   MCC1201_rgtDiagModule_HMI : GP_NetworkDiag_v1[50] := ([0].xFaulted := 1, [0].dEntryStatus := 16#0000_1000, [0].dFaultCode := 16#0000_0115, [0].dInstance := 16#0000_fdae, [1].xFaulted := 1, [1].dEntryStatus := 16#0000_1000, [1].dFaultCode := 16#0000_0115, [1].dInstance := 16#0000_3b39, [2].xConnected := 1, [2].dEntryStatus := 16#0000_4000, [2].dInstance := 16#0000_a3f5, [3].xConnected := 1, [3].dEntryStatus := 16#0000_7000, [3].dInstance := 16#0000_f5ac, [4].xConnected := 1, [4].dEntryStatus := 16#0000_7000, [4].dInstance := 16#0000_87af, [5].xFaulted := 1, [5].dEntryStatus := 16#0000_3000, [5].dFaultCode := 16#0000_0204, [5].dInstance := 16#0000_ac4a, [6].xFaulted := 1, [6].dEntryStatus := 16#0000_3000, [6].dFaultCode := 16#0000_0204, [6].dInstance := 16#0000_482b, [7].xFaulted := 1, [7].dEntryStatus := 16#0000_3000, [7].dFaultCode := 16#0000_0204, [7].dInstance := 16#0000_9886, [8].xFaulted := 1, [8].dEntryStatus := 16#0000_3000, [8].dFaultCode := 16#0000_0204, [8].dInstance := 16#0000_f085, [9].xFaulted := 1, [9].dEntryStatus := 16#0000_3000, [9].dFaultCode := 16#0000_0204, [9].dInstance := 16#0000_4058, [10].xFaulted := 1, [10].dEntryStatus := 16#0000_1000, [10].dFaultCode := 16#0000_0204, [10].dInstance := 16#0000_406f, [11].xFaulted := 1, [11].dEntryStatus := 16#0000_3000, [11].dFaultCode := 16#0000_0204, [11].dInstance := 16#0000_dc7a, [12].xConnected := 1, [12].dEntryStatus := 16#0000_4000, [12].dInstance := 16#0000_6808, [13].xConnected := 1, [13].dEntryStatus := 16#0000_4000, [13].dInstance := 16#0000_1271, [14].xConnected := 1, [14].dEntryStatus := 16#0000_4000, [14].dInstance := 16#0000_7aa0, [15].xConnected := 1, [15].dEntryStatus := 16#0000_4000, [15].dInstance := 16#0000_c3a3, [16].xConnected := 1, [16].dEntryStatus := 16#0000_4000, [16].dInstance := 16#0000_3650,
        [17].xConnected := 1, [17].dEntryStatus := 16#0000_4000, [17].dInstance := 16#0000_c67a, [18].xConnected := 1, [18].dEntryStatus := 16#0000_4000, [18].dInstance := 16#0000_cbaa, [19].xConnected := 1, [19].dEntryStatus := 16#0000_4000, [19].dInstance := 16#0000_7c6b, [20].xConnected := 1, [20].dEntryStatus := 16#0000_4000, [20].dInstance := 16#0000_b922, [21].xConnected := 1, [21].dEntryStatus := 16#0000_4000, [21].dInstance := 16#0000_0b41, [22].xConnected := 1, [22].dEntryStatus := 16#0000_4000, [22].dInstance := 16#0000_0a60, [23].xConnected := 1, [23].dEntryStatus := 16#0000_4000, [23].dInstance := 16#0000_ec63, [24].xConnected := 1, [24].dEntryStatus := 16#0000_4000, [24].dInstance := 16#0000_c43a, [25].xConnected := 1, [25].dEntryStatus := 16#0000_4000, [25].dInstance := 16#0000_ef15, [26].xConnected := 1, [26].dEntryStatus := 16#0000_4000, [26].dInstance := 16#0000_5364, [27].xConnected := 1, [27].dEntryStatus := 16#0000_4000, [27].dInstance := 16#0000_03d7, [28].xConnected := 1, [28].dEntryStatus := 16#0000_4000, [28].dInstance := 16#0000_365e, [29].xConnected := 1, [29].dEntryStatus := 16#0000_4000, [29].dInstance := 16#0000_bf29, [30].xConnected := 1, [30].dEntryStatus := 16#0000_4000, [30].dInstance := 16#0000_7fa8, [31].xConnected := 1, [31].dEntryStatus := 16#0000_4000, [31].dInstance := 16#0000_798b, [32].xConnected := 1, [32].dEntryStatus := 16#0000_4000, [32].dInstance := 16#0000_75c2, [33].xConnected := 1, [33].dEntryStatus := 16#0000_4000, [33].dInstance := 16#0000_6f7d, [34].xConnected := 1, [34].dEntryStatus := 16#0000_4000, [34].dInstance := 16#0000_332c, [35].xConnected := 1, [35].dEntryStatus := 16#0000_4000, [35].dInstance := 16#0000_e17f, [36].xConnected := 1, [36].dEntryStatus := 16#0000_4000, [36].dInstance := 16#0000_4666,
        [37].xConnected := 1, [37].dEntryStatus := 16#0000_4000, [37].dInstance := 16#0000_3411, [38].xConnected := 1, [38].xFaulted := 1, [38].dEntryStatus := 16#0000_3000, [38].dFaultCode := 16#0000_0204, [38].dInstance := 16#0000_de82, [39].xConnected := 1, [39].xFaulted := 1, [39].dEntryStatus := 16#0000_3000, [39].dFaultCode := 16#0000_0204, [39].dInstance := 16#0000_ad3d, [40].xFaulted := 1, [40].dEntryStatus := 16#0000_3000, [40].dFaultCode := 16#0000_0204, [40].dInstance := 16#0000_0f16, [41].xFaulted := 1, [41].dEntryStatus := 16#0000_1000, [41].dFaultCode := 16#0000_0204, [41].dInstance := 16#0000_0801, [42].xConnected := 1, [42].xFaulted := 1, [42].dEntryStatus := 16#0000_3000, [42].dFaultCode := 16#0000_0204, [42].dInstance := 16#0000_cb26, [43].xConnected := 1, [43].xFaulted := 1, [43].dEntryStatus := 16#0000_3000, [43].dFaultCode := 16#0000_0204, [43].dInstance := 16#0000_9dd1, [44].xConnected := 1, [44].xFaulted := 1, [44].dEntryStatus := 16#0000_3000, [44].dFaultCode := 16#0000_0204, [44].dInstance := 16#0000_2cb0, [45].xConnected := 1, [45].xFaulted := 1, [45].dEntryStatus := 16#0000_3000, [45].dFaultCode := 16#0000_0204, [45].dInstance := 16#0000_3773, [46].xConnected := 1, [46].xFaulted := 1, [46].dEntryStatus := 16#0000_3000, [46].dFaultCode := 16#0000_0204, [46].dInstance := 16#0000_0d0a, [47].xConnected := 1, [47].dEntryStatus := 16#0000_4000, [47].dInstance := 16#0000_f22b, [48].xConnected := 1, [48].dEntryStatus := 16#0000_4000, [48].dInstance := 16#0000_f6c7, [49].xConnected := 1, [49].dEntryStatus := 16#0000_4000, [49].dInstance := 16#0000_de7a); {access Read Only}
        [0]   // ETH_MCC1201_220AP1
        [11]   // MI_6CS
        [14]   // A54AZ1
        [13]   // A53AZ1
        [15]   // A55AZ1
        [17]   // A57AZ1
        [21]   // A61AZ1
        [22]   // A62AZ1
        [23]   // A63AZ1
        [24]   // A64AZ1
        [25]   // A65AZ1
        [26]   // A66AZ1
        [5]   // A152AP1
        [1]   // ETH_CULLET
        [6]   // CB_1CS
        [7]   // CB_2CS
        [8]   // CB_3CS
        [9]   // CB_4CS
        [10]   // CB_5CS
        [27]   // A67AZ1
        [28]   // A68AZ1
        [29]   // A69AZ1
        [30]   // A70AZ1
        [31]   // A71AZ1
        [32]   // A72AZ1
        [33]   // A73AZ1
        [34]   // A74AZ1
        [35]   // A75AZ1
        [36]   // A76AZ1
        [37]   // A77AZ1
        [40]   // A80AZ1
        [41]   // A81AZ1
        [4]   // Cullet_System
        [3]   // ETH_MCC1300
   MG59_000 : MESSAGE;   // PIF Operations Write current Lehr speed from N98.5 to N10:10 @ M5
        .ER   // PIF Operations Write
        MessageParameters(ServiceCode := 16#0f67, LocalElement := N98[5], ...)
   MG59_001 : MESSAGE;
   MG59_002 : MESSAGE;   // PIF Operations Write block N98:0 -> N98:3 to processor M5 N10:16 ->N10:19
        MessageParameters(ServiceCode := 16#0f67, LocalElement := N98[0], ...)
   MG59_003 : MESSAGE;
   MinorFaultBits : DINT;   // MinorFaultBits
   MS_ACCUM : ALIAS FOR N70[1];
   MS_LEHR : ALIAS FOR N60[11];
   MSEC_TRIM : ALIAS FOR N60[12];
   N : ALIAS FOR N15[80];
   N10 : DINT[128] := ([2] := 1, [3] := 32, [4] := 2050, [6] := 2, [8] := 2, [9] := 64, [10] := 4100, [12] := 4, [14] := 4, [15] := 128, [16] := 8200, [18] := 8, [20] := 8, [21] := 256, [22] := 16400, [24] := 16, [26] := 16, [27] := 512, [28] := -32736, [30] := 32, [32] := 32, [33] := 1024, [34] := 64, [35] := 1, [36] := 64, [38] := 64, [39] := 2048, [40] := 128, [41] := 2, [42] := 128, [44] := 128, [45] := 4096, [46] := 256, [47] := 4, [48] := 256, [50] := 256, [51] := 8192, [52] := 512, [53] := 8, [54] := 512, [56] := 512, [57] := 16384, [58] := 1024, [59] := 16, [60] := 1024, [62] := 1024, [63] := -32768, [64] := 1024, [65] := -32768, [66] := 1024, [68] := 1024, [69] := 16, [70] := 512, [71] := 16384, [72] := 512, [74] := 512, [75] := 8, [76] := 256, [77] := 8192, [78] := 256,
        [80] := 256, [81] := 4, [82] := 128, [83] := 4096, [84] := 128, [86] := 128, [87] := 2, [88] := 64, [89] := 2048, [90] := 64, [92] := 64, [93] := 1, [94] := 32, [95] := 1024, [96] := 32, [98] := -32736, [100] := 16, [101] := 512, [102] := 16, [104] := 16400, [106] := 8, [107] := 256, [108] := 8, [110] := 8200, [112] := 4, [113] := 128, [114] := 4, [116] := 4100, [118] := 2, [119] := 64, [120] := 2, [122] := 2050, [124] := 1, [125] := 32, [126] := 1);
   N100 : DINT[1000] := ([0] := 2683, [1] := 2683, [2] := 2683, [3] := 2683, [4] := 2683, [5] := 2683, [6] := 2683, [7] := 2683, [8] := 2683, [9] := 2683, [10] := 2683, [11] := 2683, [12] := 2683, [13] := 2683, [14] := 2683, [15] := 2683, [16] := 2683, [17] := 2683, [18] := 2683, [19] := 2683, [20] := 2683, [21] := 2683, [22] := 2683, [23] := 2683, [24] := 2683, [25] := 2683, [26] := 2683, [27] := 2683, [28] := 2683, [29] := 2683, [30] := 2683, [31] := 2683, [32] := 2683, [33] := 2683, [34] := 2683, [35] := 2683, [36] := 2683, [37] := 2683, [38] := 2683, [39] := 2683, [40] := 2683, [41] := 2683, [42] := 2683, [43] := 2683, [44] := 2683, [45] := 2683, [46] := 2683, [47] := 2683, [48] := 2683, [49] := 2683, [50] := 2683, [51] := 2683, [52] := 2683, [53] := 2683, [54] := 2683, [55] := 2683, [56] := 2683, [57] := 2683, [58] := 2683, [59] := 2683,
        [60] := 2683, [61] := 2683, [62] := 2683, [63] := 2683, [64] := 2683, [65] := 2683, [66] := 2683, [67] := 2683, [68] := 2683, [69] := 2683, [70] := 2683, [71] := 2683, [72] := 2683, [73] := 2683, [74] := 2683, [75] := 2683, [76] := 2683, [77] := 2683, [78] := 2683, [79] := 2683, [80] := 2683, [81] := 2683, [82] := 2683, [83] := 2683, [84] := 2683, [85] := 2683, [86] := 2683, [87] := 2683, [88] := 2683, [89] := 2683, [90] := 2683, [91] := 2683, [92] := 2683, [93] := 2683, [94] := 2683, [95] := 2683, [96] := 2683, [97] := 2683, [98] := 2683, [99] := 2683, [100] := 2683, [101] := 2683, [102] := 2683, [103] := 2683, [104] := 2683, [105] := 2683, [106] := 2683, [107] := 2683, [108] := 2683, [109] := 2683, [110] := 2683, [111] := 2683, [112] := 2683, [113] := 2683, [114] := 2683, [115] := 2683, [116] := 2683, [117] := 2683, [118] := 2683, [119] := 2683,
        [120] := 2683, [121] := 2683, [122] := 2683, [123] := 2683, [124] := 2683, [125] := 2683, [126] := 2683, [127] := 2683, [128] := 2683, [129] := 2683, [130] := 2683, [131] := 2683, [132] := 2683, [133] := 2683, [134] := 2683, [135] := 2683, [136] := 2683, [137] := 2683, [138] := 2683, [139] := 2683, [140] := 2683, [141] := 2683, [142] := 2683, [143] := 2683, [144] := 2683, [145] := 2683, [146] := 2683, [147] := 2683, [148] := 2683, [149] := 2683, [150] := 2683, [151] := 2683, [152] := 2683, [153] := 2683, [154] := 2683, [155] := 2683, [156] := 2683, [157] := 2683, [158] := 2683, [159] := 2683, [160] := 2683, [161] := 2683, [162] := 2683, [163] := 2683, [164] := 2683, [165] := 2683, [166] := 2683, [167] := 2683, [168] := 2683, [169] := 2683, [170] := 2683, [171] := 2683, [172] := 2683, [173] := 2683, [174] := 2683, [175] := 2683, [176] := 2683, [177] := 2683, [178] := 2683, [179] := 2683,
        [180] := 2683, [181] := 2683, [182] := 2683, [183] := 2683, [184] := 2683, [185] := 2683, [186] := 2683, [187] := 2683, [188] := 2683, [189] := 2683, [190] := 2683, [191] := 2683, [192] := 2683, [193] := 2683, [194] := 2683, [195] := 2683, [196] := 2683, [197] := 2683, [198] := 2683, [199] := 2683, [200] := 2683, [201] := 2683, [202] := 2683, [203] := 2683, [204] := 2683, [205] := 2683, [206] := 2683, [207] := 2683, [208] := 2683, [209] := 2683, [210] := 2683, [211] := 2683, [212] := 2683, [213] := 2683, [214] := 2683, [215] := 2683, [216] := 2683, [217] := 2683, [218] := 2683, [219] := 2683, [220] := 2683, [221] := 2683, [222] := 2683, [223] := 2683, [224] := 2683, [225] := 2683, [226] := 2683, [227] := 2683, [228] := 2683, [229] := 2683, [230] := 2683, [231] := 2683, [232] := 2683, [233] := 2683, [234] := 2683, [235] := 2683, [236] := 2683, [237] := 2683, [238] := 2683, [239] := 2683,
        [240] := 2683, [241] := 2683, [242] := 2683, [243] := 2683, [244] := 2683, [245] := 2683, [246] := 2683, [247] := 2683, [248] := 2683, [249] := 2683, [250] := 2683, [251] := 2683, [252] := 2683, [253] := 2683, [254] := 2683, [255] := 2683, [256] := 2683, [257] := 2683, [258] := 2683, [259] := 2683, [260] := 2683, [261] := 2683, [262] := 2683, [263] := 2683, [264] := 2683, [265] := 2683, [266] := 2683, [267] := 2683, [268] := 2683, [269] := 2683, [270] := 2683, [271] := 2683, [272] := 2683, [273] := 2683, [274] := 2683, [275] := 2683, [276] := 2683, [277] := 2683, [278] := 2683, [279] := 2683, [280] := 2683, [281] := 2683, [282] := 2683, [283] := 2683, [284] := 2683, [285] := 2683, [286] := 2683, [287] := 2683, [288] := 2683, [289] := 2683, [290] := 2683, [291] := 2683, [292] := 2683, [293] := 2683, [294] := 2683, [295] := 2683, [296] := 2683, [297] := 2683, [298] := 2683, [299] := 2683,
        [300] := 2683, [301] := 2683, [302] := 2683, [303] := 2683, [304] := 2686, [305] := 2676, [306] := 2681, [307] := 2679, [308] := 2686, [309] := 2679, [310] := 2691, [311] := 2679, [312] := 2681, [313] := 2681, [314] := 2688, [315] := 2688, [316] := 2686, [317] := 2683, [318] := 2686, [319] := 2693, [320] := 2787, [321] := 2794, [322] := 2787, [323] := 2785, [324] := 2792, [325] := 2794, [326] := 2792, [327] := 2785, [328] := 2783, [329] := 2787, [330] := 2797, [331] := 2792, [332] := 2799, [333] := 2792, [334] := 2818, [335] := 2790, [336] := 2792, [337] := 2783, [338] := 2783, [339] := 2792, [340] := 2794, [341] := 2797, [342] := 2792, [343] := 2794, [344] := 2787, [345] := 2787, [346] := 2783, [347] := 2785, [348] := 2797, [349] := 2794, [350] := 2787, [351] := 2787, [352] := 2780, [353] := 2790, [354] := 2787, [355] := 2794, [356] := 2792, [357] := 2783, [358] := 2787, [359] := 2783,
        [360] := 2809, [361] := 2806, [362] := 2828, [363] := 2813, [364] := 2804, [365] := 2794, [366] := 2790, [367] := 2794, [368] := 2794, [369] := 2790, [370] := 2794, [371] := 2787, [372] := 2797, [373] := 2797, [374] := 2792, [375] := 2799, [376] := 2792, [377] := 2792, [378] := 2787, [379] := 2785, [380] := 2802, [381] := 2799, [382] := 2794, [383] := 2792, [384] := 2794, [385] := 2787, [386] := 2797, [387] := 2797, [388] := 2794, [389] := 2787, [390] := 2794, [391] := 2787, [392] := 2792, [393] := 2790, [394] := 2797, [395] := 2794, [396] := 2794, [397] := 2787, [398] := 2794, [399] := 2787, [400] := 2799, [401] := 2799, [402] := 2797, [403] := 2794, [404] := 2790, [405] := 2787, [406] := 2787, [407] := 2818, [408] := 2811, [409] := 2806, [410] := 2799, [411] := 2790, [412] := 2792, [413] := 2785, [414] := 2787, [415] := 2792, [416] := 2799, [417] := 2802, [418] := 2797, [419] := 2806,
        [420] := 2802, [421] := 2792, [422] := 2799, [423] := 2804, [424] := 2813, [425] := 2792, [426] := 2828, [427] := 2809, [428] := 2783, [429] := 2832, [430] := 2806, [431] := 2811, [432] := 2804, [433] := 2804, [434] := 2813, [435] := 2804, [436] := 2809, [437] := 2816, [438] := 2816, [439] := 2811, [440] := 2811, [441] := 2806, [442] := 2828, [443] := 2792, [444] := 2816, [445] := 2806, [446] := 2797, [447] := 2816, [448] := 2799, [449] := 2799, [450] := 2811, [451] := 2799, [452] := 2797, [453] := 2797, [454] := 2802, [455] := 2778, [456] := 2776, [457] := 2783, [458] := 2792, [459] := 2769, [460] := 2776, [461] := 2776, [462] := 2769, [463] := 2771, [464] := 2769, [465] := 2769, [466] := 2773, [467] := 2769, [468] := 2776, [469] := 2764, [470] := 2766, [471] := 2683, [472] := 2686, [473] := 2702, [474] := 2691, [475] := 2705, [476] := 2688, [477] := 2698, [478] := 2700, [479] := 2686,
        [480] := 2702, [481] := 2683, [482] := 2691, [483] := 2695, [484] := 2688, [485] := 2712, [486] := 2691, [487] := 2700, [488] := 2698, [489] := 2695, [490] := 2700, [491] := 2691, [492] := 2693, [493] := 2693, [494] := 2693, [495] := 2707, [496] := 2695, [497] := 2693, [498] := 2693, [499] := 2683, [500] := 2681, [501] := 2688, [502] := 2691, [503] := 2688, [504] := 2691, [505] := 2681, [506] := 2681, [507] := 2688, [508] := 2686, [509] := 2693, [510] := 2681, [511] := 2676, [512] := 2674, [513] := 2683, [514] := 2693, [515] := 2693, [516] := 2681, [517] := 2683, [518] := 2681, [519] := 2693, [520] := 2688, [521] := 2683, [522] := 2681, [523] := 2676, [524] := 2679, [525] := 2688, [526] := 2693, [527] := 2681, [528] := 2679, [529] := 2679, [530] := 2695, [531] := 2686, [532] := 2679, [533] := 2676, [534] := 2679, [535] := 2688, [536] := 2686, [537] := 2688, [538] := 2679, [539] := 2679,
        [540] := 2676, [541] := 2686, [542] := 2686, [543] := 2676, [544] := 2676, [545] := 2674, [546] := 2681, [547] := 2691, [548] := 2688, [549] := 2688, [550] := 2693, [551] := 2705, [552] := 2681, [553] := 2681, [554] := 2719, [555] := 2688, [556] := 2695, [557] := 2702, [558] := 2688, [559] := 2688, [560] := 2700, [561] := 2700, [562] := 2679, [563] := 2681, [564] := 2688, [565] := 2681, [566] := 2681, [567] := 2686, [568] := 2681, [569] := 2683, [570] := 2693, [571] := 2686, [572] := 2676, [573] := 2679, [574] := 2681, [575] := 2683, [576] := 2686, [577] := 2693, [578] := 2679, [579] := 2679, [580] := 2681, [581] := 2679, [582] := 2688, [583] := 2683, [584] := 2674, [585] := 2681, [586] := 2676, [587] := 2679, [588] := 2681, [589] := 2686, [590] := 2698, [591] := 2683, [592] := 2683, [593] := 2679, [594] := 2686, [595] := 2771, [596] := 2780, [597] := 2780, [598] := 2778, [599] := 2776,
        [600] := 2773, [601] := 2780, [602] := 2771, [603] := 2780, [604] := 2785, [605] := 2778, [606] := 2773, [607] := 2773, [608] := 2783, [609] := 2769, [610] := 2780, [611] := 2780, [612] := 2773, [613] := 2780, [614] := 2771, [615] := 2778, [616] := 2769, [617] := 2769, [618] := 2790, [619] := 2776, [620] := 2783, [621] := 2771, [622] := 2778, [623] := 2773, [624] := 2776, [625] := 2780, [626] := 2773, [627] := 2790, [628] := 2769, [629] := 2785, [630] := 2780, [631] := 2773, [632] := 2787, [633] := 2778, [634] := 2783, [635] := 2776, [636] := 2776, [637] := 2776, [638] := 2783, [639] := 2787, [640] := 2776, [641] := 2783, [642] := 2776, [643] := 2773, [644] := 2783, [645] := 2769, [646] := 2776, [647] := 2776, [648] := 2773, [649] := 2769, [650] := 2778, [651] := 2780, [652] := 2773, [653] := 2783, [654] := 2773, [655] := 2773, [656] := 2773, [657] := 2776, [658] := 2785, [659] := 2778,
        [660] := 2785, [661] := 2771, [662] := 2776, [663] := 2778, [664] := 2776, [665] := 2778, [666] := 2771, [667] := 2787, [668] := 2773, [669] := 2783, [670] := 2787, [671] := 2773, [672] := 2773, [673] := 2771, [674] := 2776, [675] := 2778, [676] := 2790, [677] := 2766, [678] := 2787, [679] := 2785, [680] := 2780, [681] := 2785, [682] := 2771, [683] := 2778, [684] := 2771, [685] := 2780, [686] := 2771, [687] := 2766, [688] := 2776, [689] := 2776, [690] := 2769, [691] := 2773, [692] := 2773, [693] := 2771, [694] := 2776, [695] := 2778, [696] := 2766, [697] := 2771, [698] := 2783, [699] := 2761, [700] := 2766, [701] := 2778, [702] := 2776, [703] := 2776, [704] := 2757, [705] := 2757, [706] := 2759, [707] := 2750, [708] := 2778, [709] := 2776, [710] := 2764, [711] := 2759, [712] := 2757, [713] := 2766, [714] := 2757, [715] := 2757, [716] := 2757, [717] := 2676, [718] := 2683, [719] := 2691,
        [720] := 2691, [721] := 2686, [722] := 2681, [723] := 2688, [724] := 2679, [725] := 2688, [726] := 2691, [727] := 2693, [728] := 2683, [729] := 2681, [730] := 2683, [731] := 2681, [732] := 2693, [733] := 2693, [734] := 2695, [735] := 2698, [736] := 2693, [737] := 2698, [738] := 2693, [739] := 2693, [740] := 2691, [741] := 2702, [742] := 2695, [743] := 2712, [744] := 2693, [745] := 2717, [746] := 2702, [747] := 2709, [748] := 2707, [749] := 2695, [750] := 2679, [751] := 2731, [752] := 2783, [753] := 2794, [754] := 2785, [755] := 2783, [756] := 2794, [757] := 2792, [758] := 2787, [759] := 2787, [760] := 2797, [761] := 2787, [762] := 2785, [763] := 2792, [764] := 2787, [765] := 2787, [766] := 2806, [767] := 2780, [768] := 2783, [769] := 2794, [770] := 2783, [771] := 2783, [772] := 2794, [773] := 2790, [774] := 2783, [775] := 2790, [776] := 2794, [777] := 2785, [778] := 2785, [779] := 2790,
        [780] := 2792, [781] := 2783, [782] := 2790, [783] := 2790, [784] := 2778, [785] := 2787, [786] := 2790, [787] := 2787, [788] := 2783, [789] := 2802, [790] := 2787, [791] := 2794, [792] := 2790, [793] := 2773, [794] := 2776, [795] := 2778, [796] := 2783, [797] := 2776, [798] := 2787, [799] := 2776, [800] := 2787, [801] := 2776, [802] := 2787, [803] := 2769, [804] := 2780, [805] := 2771, [806] := 2787, [807] := 2773, [808] := 2785, [809] := 2771, [810] := 2785, [811] := 2776, [812] := 2778, [813] := 2773, [814] := 2780, [815] := 2771, [816] := 2783, [817] := 2778, [818] := 2780, [819] := 2790, [820] := 2778, [821] := 2785, [822] := 2771, [823] := 2785, [824] := 2776, [825] := 2787, [826] := 2776, [827] := 2787, [828] := 2773, [829] := 2780, [830] := 2773, [831] := 2780, [832] := 2783, [833] := 2785, [834] := 2769, [835] := 2787, [836] := 2766, [837] := 2778, [838] := 2778, [839] := 2776,
        [840] := 2787, [841] := 2776, [842] := 2780, [843] := 2778, [844] := 2773, [845] := 2778, [846] := 2776, [847] := 2780, [848] := 2783, [849] := 2766, [850] := 2787, [851] := 2773, [852] := 2776, [853] := 2773, [854] := 2780, [855] := 2771, [856] := 2778, [857] := 2771, [858] := 2776, [859] := 2780, [860] := 2785, [861] := 2776, [862] := 2783, [863] := 2776, [864] := 2780, [865] := 2766, [866] := 2776, [867] := 432, [868] := 432, [869] := 2806, [870] := 2797, [871] := 2773, [872] := 531, [873] := 2776, [874] := 2792, [875] := 2790, [876] := 2783, [877] := 2778, [878] := 2780, [879] := 2776, [880] := 2780, [881] := 2771, [882] := 2769, [883] := 2778, [884] := 2780, [885] := 2769, [886] := 2785, [887] := 2776, [888] := 2790, [889] := 2769, [890] := 2785, [891] := 2773, [892] := 2785, [893] := 2776, [894] := 2783, [895] := 2780, [896] := 2785, [897] := 2773, [898] := 2785, [899] := 2778,
        [900] := 2679, [901] := 2691, [902] := 2688, [903] := 2679, [904] := 2676, [905] := 2679, [906] := 2676, [907] := 2679, [908] := 2679, [909] := 2688, [910] := 2691, [911] := 2679, [912] := 2674, [913] := 2681, [914] := 2674, [915] := 2679, [916] := 2681, [917] := 2686, [918] := 2688, [919] := 2693, [920] := 2686, [921] := 2679, [922] := 2674, [923] := 2674, [924] := 2674, [925] := 2743, [926] := 2773, [927] := 2787, [928] := 2776, [929] := 2790, [930] := 2776, [931] := 2776, [932] := 2778, [933] := 2778, [934] := 2771, [935] := 2783, [936] := 2771, [937] := 2780, [938] := 2773, [939] := 2778, [940] := 2769, [941] := 2780, [942] := 2776, [943] := 2776, [944] := 2776, [945] := 2773, [946] := 2785, [947] := 2778, [948] := 2776, [949] := 2776, [950] := 2773, [951] := 2776, [952] := 2778, [953] := 2773, [954] := 2785, [955] := 2771, [956] := 2790, [957] := 2776, [958] := 2764, [959] := 2769,
        [960] := 2769, [961] := 2766, [962] := 2759, [963] := 2761, [964] := 2764, [965] := 2761, [966] := 2776, [967] := 2783, [968] := 2766, [969] := 2757, [970] := 2752, [971] := 2752, [972] := 2754, [973] := 2754, [974] := 2754, [975] := 2750, [976] := 2747, [977] := 2745, [978] := 2754, [979] := 2752, [980] := 2766, [981] := 2761, [982] := 2761, [983] := 2764, [984] := 2764, [985] := 2757, [986] := 2752, [987] := 2766, [988] := 2759, [989] := 2759, [990] := 2771, [991] := 2752, [992] := 2752, [993] := 2752, [994] := 2750, [995] := 2773, [996] := 2771, [997] := 2757, [998] := 2759, [999] := 2754);
   N11 : DINT[1000];
        [0]   // Scanner 5 Traking File
   N11_HOST : INT[1000]; {produced}
   N12 : DINT[1000];
   N124 : DINT[414] := ([0] := 3269, [250] := 2, [254] := 254, [350] := 28673, [351] := 256, [352] := -28665, [383] := 256, [384] := -28671);
   N125 : DINT[414] := ([5] := 100, [6] := 5064, [127] := 100, [128] := 3000, [135] := 100, [136] := 3000, [143] := 100, [144] := 3000, [151] := 100, [152] := 3000, [159] := 100, [160] := 1816, [167] := 100, [168] := 1816, [351] := 7, [352] := 4096, [353] := 148, [355] := 2, [356] := 1, [382] := 28673, [383] := 263, [384] := 4096, [385] := 148, [387] := 2, [388] := 1);
        [160]   // Washer Sponge Upper Roll Speed Ref Via Device Net
        [168]   // Washer Sponge Lower Roll Speed Ref Via Device Net
   N126 : DINT[103] := ([0] := 24, [1] := 27, [2] := 28, [3] := 29, [4] := 73, [5] := 74, [6] := 75, [7] := 76, [8] := 7, [9] := 8, [10] := 158, [11] := 159, [12] := 40, [13] := 91, [14] := 122, [15] := 123, [16] := 124, [17] := 114, [18] := 115, [19] := 116, [20] := 19, [21] := 21, [22] := 10, [23] := 38, [24] := 36, [25] := 5, [26] := 6, [27] := 94, [28] := 95, [29] := 96, [30] := 97, [31] := 98, [32] := 99, [33] := 100, [34] := 92, [35] := 93, [36] := 192, [37] := 193, [38] := 85, [39] := 37, [40] := 57, [50] := 60, [51] := 147, [52] := 170, [53] := 171, [54] := 65, [55] := 66, [56] := 1, [57] := 54, [58] := 23, [59] := 162, [60] := 163, [61] := 2, [62] := 3, [63] := 53, [64] := 70, [65] := 4, [66] := 86, [67] := 87, [68] := 88,
        [69] := 89, [70] := 143, [71] := 144, [72] := 145, [73] := 146, [74] := 173, [75] := 59, [76] := 55, [77] := 62, [78] := 141, [79] := 142, [101] := 1, [102] := 7);
        [101]   // DEVICENET Number of Drives ** channel a **
        [102]   // DEVICENET Number of Drives ** channel b **
   N127 : DINT[997] := ([0] := 1000, [36] := 6000, [96] := 100, [108] := 300, [168] := 27, [204] := 27, [240] := 90, [252] := 12, [264] := 2, [276] := 4710, [288] := 6144, [300] := 6, [312] := 12, [324] := 1, [336] := 1, [348] := 1, [360] := 1, [372] := 1, [384] := 1, [396] := 5, [408] := 5, [444] := 300, [456] := 3, [612] := 460, [624] := 84, [636] := 370, [648] := 19070, [672] := 3582, [684] := 871, [696] := 532, [708] := 354, [720] := 803, [732] := 858, [744] := 512, [756] := 5902, [768] := 54, [780] := 10, [792] := 10, [804] := 2, [816] := 10, [828] := 2, [840] := 1, [852] := 2, [888] := 1, [912] := 83, [924] := 12, [936] := 6, [948] := 8, [990] := 1, [994] := 1, [996] := 1);